// TIA Portal project "Sistema_de_silos" (V16) (continued)
REGION Network 7: Acionamento do Damper / Logica de segurança
   // O ideal é ter o feedback do motor (transportador)
   RUNG wire#powerrail
      Contact( #iCmdAbasteceSilo )
      I_Contact( #iSensorMaximo )
      wire#w1
      Contact( #iSensorDamper01 )
      Contact( #iSensorDamper02 )
      wire#w2
      I_Contact( #Falha_SensoresNivel )
      I_Contact( #Falha_TimeOut_Desabastecimento )
      I_Contact( #iEmg )
      I_Contact( #iCodinicial )
      Coil( #oLigarDumper )
   END_RUNG
   RUNG wire#w1
      Contact( #oLigarDumper )
   END_RUNG wire#w2
   RUNG wire#powerrail
      Contact( #iManual )
      Contact( #btnLigaDumper )
      I_Contact( #"Status Silo - Maximo" )
      Contact( #oLigarTransportador )
      I_Contact( #protecao_damper )
   END_RUNG wire#w2
   // the same network as SCL:
   #oLigarDumper := ((#iCmdAbasteceSilo AND NOT #iSensorMaximo AND ((#iSensorDamper01 AND #iSensorDamper02) OR #oLigarDumper)) OR (#iManual AND #btnLigaDumper AND NOT #"Status Silo - Maximo" AND #oLigarTransportador AND NOT #protecao_damper)) AND NOT #Falha_SensoresNivel AND NOT #Falha_TimeOut_Desabastecimento AND NOT #iEmg AND NOT #iCodinicial;
END_REGION

REGION Network 8: Liga Transportador
   RUNG wire#powerrail
      Contact( #status_damper )
      Contact( #iAutomatico )
      wire#w1
      I_Contact( #Falha_SensoresNivel )
      I_Contact( #Falha_TimeOut_Desabastecimento )
      I_Contact( #iEmg )
      Coil( #oLigarTransportador )
   END_RUNG
   RUNG wire#powerrail
      Contact( #iManual )
      Contact( #btnLigaTransportador )
   END_RUNG wire#w1
   // the same network as SCL:
   #oLigarTransportador := ((#status_damper AND #iAutomatico) OR (#iManual AND #btnLigaTransportador)) AND NOT #Falha_SensoresNivel AND NOT #Falha_TimeOut_Desabastecimento AND NOT #iEmg;
END_REGION

REGION Network 9: Silo Principal - Reserva do produto
   RUNG wire#powerrail
      Contact( #iSensorMinimo )
      wire#w1
      I_Contact( #iSensorMaximo )
      Coil( #"Status Silo - Minimo" )
   END_RUNG
   RUNG wire#w1
      Contact( #iSensorMaximo )
      Coil( #"Status Silo - Maximo" )
   END_RUNG
   RUNG wire#powerrail
      I_Contact( #iSensorMinimo )
      I_Contact( #iSensorMaximo )
      Coil( #"Status Silo - Desabastecido" )
   END_RUNG
   // the same network as SCL:
   #"Status Silo - Minimo" := #iSensorMinimo AND NOT #iSensorMaximo;
   #"Status Silo - Maximo" := #iSensorMinimo AND #iSensorMaximo;
   #"Status Silo - Desabastecido" := NOT #iSensorMinimo AND NOT #iSensorMaximo;
END_REGION

REGION Network 10: Falha dos Sensores de Nivel
   RUNG wire#powerrail
      Contact( #iSensorMaximo )
      I_Contact( #iSensorMinimo )
      S_Coil( #Falha_SensoresNivel )
   END_RUNG
   // the same network as SCL:
   IF #iSensorMaximo AND NOT #iSensorMinimo THEN #Falha_SensoresNivel := TRUE; END_IF;
END_REGION

REGION Network 11: Memoria Auxilar de Erro - Falha de desabastecimento
   RUNG wire#powerrail
      Contact( #"Status Silo - Minimo" )
      Contact( #oAbrirValvula )
      I_Contact( #"Status Silo - Maximo" )
      S_Coil( "DB_Geral".Memoria_Auxiliar_Erro_Silo_1 )
   END_RUNG
   RUNG wire#powerrail
      Contact( #"Status Silo - Desabastecido" )
      R_Coil( "DB_Geral".Memoria_Auxiliar_Erro_Silo_1 )
   END_RUNG
   // the same network as SCL:
   IF #"Status Silo - Minimo" AND #oAbrirValvula AND NOT #"Status Silo - Maximo" THEN
       "DB_Geral".Memoria_Auxiliar_Erro_Silo_1 := TRUE;
   END_IF;
   IF #"Status Silo - Desabastecido" THEN "DB_Geral".Memoria_Auxiliar_Erro_Silo_1 := FALSE; END_IF;
END_REGION

REGION Network 12: Falha de Desabastecimento
   "IEC_Timer_0_DB_TON_TempoErro".TON(IN := "DB_Geral".Memoria_Auxiliar_Erro_Silo_1,
                           PT := "DB_Geral".Time_TempoErro_1);
   IF "IEC_Timer_0_DB_TON_TempoErro".Q THEN #Falha_TimeOut_Desabastecimento := TRUE; END_IF;
END_REGION

REGION Network 13: Reset - Falhas
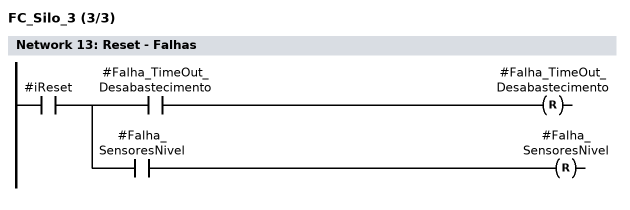
   RUNG wire#powerrail
      Contact( #iReset )
      wire#w1
      Contact( #Falha_TimeOut_Desabastecimento )
      R_Coil( #Falha_TimeOut_Desabastecimento )
   END_RUNG
   RUNG wire#w1
      Contact( #Falha_SensoresNivel )
      R_Coil( #Falha_SensoresNivel )
   END_RUNG
   // the same network as SCL:
   IF #iReset AND #Falha_TimeOut_Desabastecimento THEN #Falha_TimeOut_Desabastecimento := FALSE; END_IF;
   IF #iReset AND #Falha_SensoresNivel THEN #Falha_SensoresNivel := FALSE; END_IF;
END_REGION
END_FUNCTION

FUNCTION "FC_estado_Silos" : Void   // FC8, LAD
{ S7_Optimized_Access := 'TRUE' }
VERSION : 0.1
BEGIN

REGION Network 1
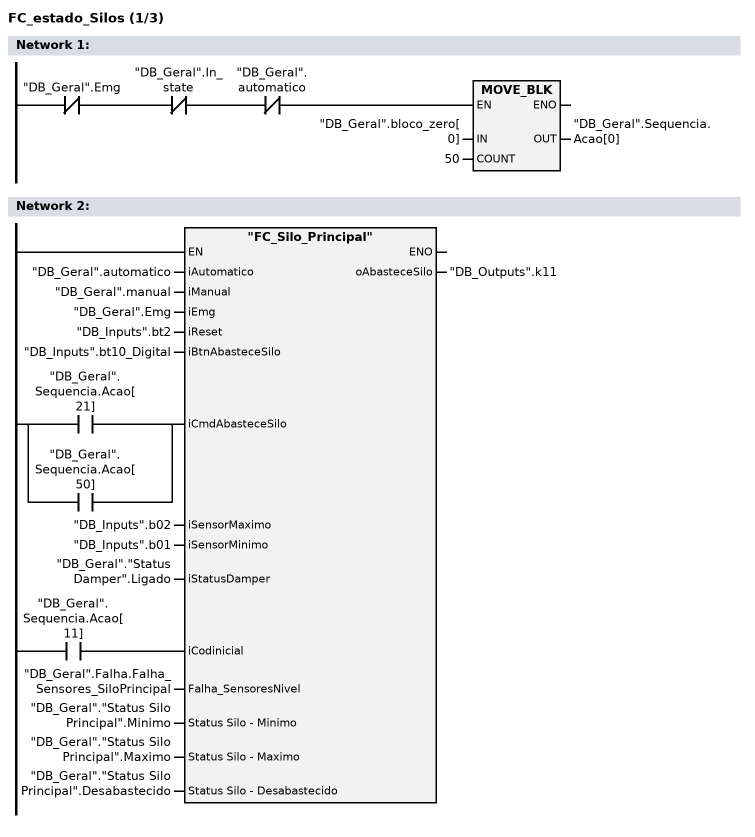
   IF NOT "DB_Geral".Emg AND NOT "DB_Geral".In_state AND NOT "DB_Geral".automatico THEN
       MOVE_BLK(IN := "DB_Geral".bloco_zero[0], COUNT := 50, OUT => "DB_Geral".Sequencia.Acao[0]);
   END_IF;
END_REGION

REGION Network 2
   RUNG wire#powerrail
      "FC_Silo_Principal"(iCmdAbasteceSilo := wire#w1, iCodinicial := wire#w2, iAutomatico := "DB_Geral".automatico, iManual := "DB_Geral".manual, iEmg := "DB_Geral".Emg, iReset := "DB_Inputs".bt2, iBtnAbasteceSilo := "DB_Inputs".bt10_Digital, iSensorMaximo := "DB_Inputs".b02, iSensorMinimo := "DB_Inputs".b01, iStatusDamper := "DB_Geral"."Status Damper".Ligado, Falha_SensoresNivel := "DB_Geral".Falha.Falha_Sensores_SiloPrincipal, "Status Silo - Minimo" := "DB_Geral"."Status Silo Principal".Minimo, "Status Silo - Maximo" := "DB_Geral"."Status Silo Principal".Maximo, "Status Silo - Desabastecido" := "DB_Geral"."Status Silo Principal".Desabastecido, oAbasteceSilo => "DB_Outputs".k11)
   END_RUNG
   RUNG wire#powerrail
      Contact( "DB_Geral".Sequencia.Acao[21] )
   END_RUNG wire#w1
   RUNG wire#powerrail
      Contact( "DB_Geral".Sequencia.Acao[50] )
   END_RUNG wire#w1
   RUNG wire#powerrail
      Contact( "DB_Geral".Sequencia.Acao[11] )
   END_RUNG wire#w2
   // the same network as SCL:
   "FC_Silo_Principal"(iAutomatico := "DB_Geral".automatico,
                       iManual := "DB_Geral".manual,
                       iEmg := "DB_Geral".Emg,
                       iReset := "DB_Inputs".bt2,
                       iBtnAbasteceSilo := "DB_Inputs".bt10_Digital,
                       iCmdAbasteceSilo := "DB_Geral".Sequencia.Acao[21] OR "DB_Geral".Sequencia.Acao[50],
                       iSensorMaximo := "DB_Inputs".b02,
                       iSensorMinimo := "DB_Inputs".b01,
                       iStatusDamper := "DB_Geral"."Status Damper".Ligado,
                       iCodinicial := "DB_Geral".Sequencia.Acao[11],
                       Falha_SensoresNivel := "DB_Geral".Falha.Falha_Sensores_SiloPrincipal,
                       "Status Silo - Minimo" := "DB_Geral"."Status Silo Principal".Minimo,
                       "Status Silo - Maximo" := "DB_Geral"."Status Silo Principal".Maximo,
                       "Status Silo - Desabastecido" := "DB_Geral"."Status Silo Principal".Desabastecido,
                       oAbasteceSilo => "DB_Outputs".k11);
END_REGION

REGION Network 3
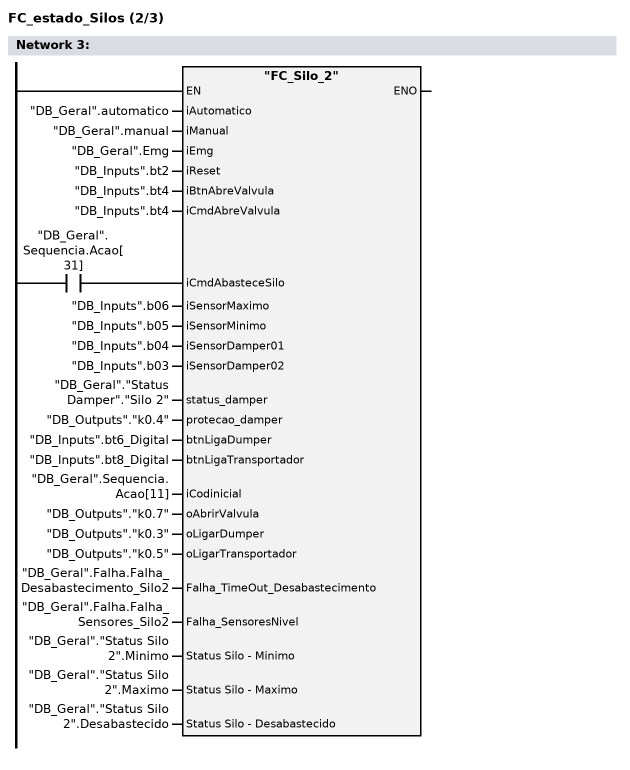
   RUNG wire#powerrail
      "FC_Silo_2"(iCmdAbasteceSilo := wire#w1, iAutomatico := "DB_Geral".automatico, iManual := "DB_Geral".manual, iEmg := "DB_Geral".Emg, iReset := "DB_Inputs".bt2, iBtnAbreValvula := "DB_Inputs".bt4, iCmdAbreValvula := "DB_Inputs".bt4, iSensorMaximo := "DB_Inputs".b06, iSensorMinimo := "DB_Inputs".b05, iSensorDamper01 := "DB_Inputs".b04, iSensorDamper02 := "DB_Inputs".b03, status_damper := "DB_Geral"."Status Damper"."Silo 2", protecao_damper := "DB_Outputs"."k0.4", btnLigaDumper := "DB_Inputs".bt6_Digital, btnLigaTransportador := "DB_Inputs".bt8_Digital, iCodinicial := "DB_Geral".Sequencia.Acao[11], oAbrirValvula := "DB_Outputs"."k0.7", oLigarDumper := "DB_Outputs"."k0.3", oLigarTransportador := "DB_Outputs"."k0.5", Falha_TimeOut_Desabastecimento := "DB_Geral".Falha.Falha_Desabastecimento_Silo2, Falha_SensoresNivel := "DB_Geral".Falha.Falha_Sensores_Silo2, "Status Silo - Minimo" := "DB_Geral"."Status Silo 2".Minimo, "Status Silo - Maximo" := "DB_Geral"."Status Silo 2".Maximo, "Status Silo - Desabastecido" := "DB_Geral"."Status Silo 2".Desabastecido)
   END_RUNG
   RUNG wire#powerrail
      Contact( "DB_Geral".Sequencia.Acao[31] )
   END_RUNG wire#w1
   // the same network as SCL:
   "FC_Silo_2"(iAutomatico := "DB_Geral".automatico,
               iManual := "DB_Geral".manual,
               iEmg := "DB_Geral".Emg,
               iReset := "DB_Inputs".bt2,
               iBtnAbreValvula := "DB_Inputs".bt4,
               iCmdAbreValvula := "DB_Inputs".bt4,
               iCmdAbasteceSilo := "DB_Geral".Sequencia.Acao[31],
               iSensorMaximo := "DB_Inputs".b06,
               iSensorMinimo := "DB_Inputs".b05,
               iSensorDamper01 := "DB_Inputs".b04,
               iSensorDamper02 := "DB_Inputs".b03,
               status_damper := "DB_Geral"."Status Damper"."Silo 2",
               protecao_damper := "DB_Outputs"."k0.4",
               btnLigaDumper := "DB_Inputs".bt6_Digital,
               btnLigaTransportador := "DB_Inputs".bt8_Digital,
               iCodinicial := "DB_Geral".Sequencia.Acao[11],
               oAbrirValvula := "DB_Outputs"."k0.7",
               oLigarDumper := "DB_Outputs"."k0.3",
               oLigarTransportador := "DB_Outputs"."k0.5",
               Falha_TimeOut_Desabastecimento := "DB_Geral".Falha.Falha_Desabastecimento_Silo2,
               Falha_SensoresNivel := "DB_Geral".Falha.Falha_Sensores_Silo2,
               "Status Silo - Minimo" := "DB_Geral"."Status Silo 2".Minimo,
               "Status Silo - Maximo" := "DB_Geral"."Status Silo 2".Maximo,
               "Status Silo - Desabastecido" := "DB_Geral"."Status Silo 2".Desabastecido);
END_REGION

REGION Network 4
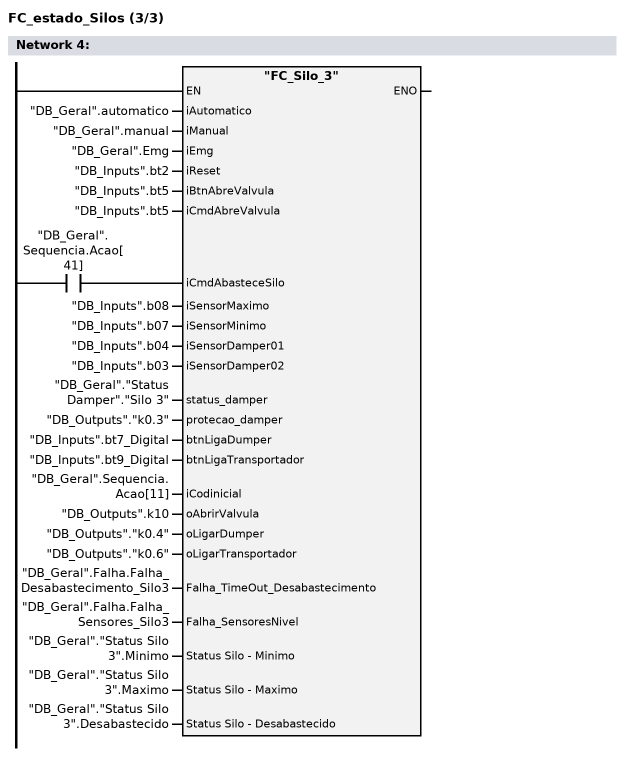
   RUNG wire#powerrail
      "FC_Silo_3"(iCmdAbasteceSilo := wire#w1, iAutomatico := "DB_Geral".automatico, iManual := "DB_Geral".manual, iEmg := "DB_Geral".Emg, iReset := "DB_Inputs".bt2, iBtnAbreValvula := "DB_Inputs".bt5, iCmdAbreValvula := "DB_Inputs".bt5, iSensorMaximo := "DB_Inputs".b08, iSensorMinimo := "DB_Inputs".b07, iSensorDamper01 := "DB_Inputs".b04, iSensorDamper02 := "DB_Inputs".b03, status_damper := "DB_Geral"."Status Damper"."Silo 3", protecao_damper := "DB_Outputs"."k0.3", btnLigaDumper := "DB_Inputs".bt7_Digital, btnLigaTransportador := "DB_Inputs".bt9_Digital, iCodinicial := "DB_Geral".Sequencia.Acao[11], oAbrirValvula := "DB_Outputs".k10, oLigarDumper := "DB_Outputs"."k0.4", oLigarTransportador := "DB_Outputs"."k0.6", Falha_TimeOut_Desabastecimento := "DB_Geral".Falha.Falha_Desabastecimento_Silo3, Falha_SensoresNivel := "DB_Geral".Falha.Falha_Sensores_Silo3, "Status Silo - Minimo" := "DB_Geral"."Status Silo 3".Minimo, "Status Silo - Maximo" := "DB_Geral"."Status Silo 3".Maximo, "Status Silo - Desabastecido" := "DB_Geral"."Status Silo 3".Desabastecido)
   END_RUNG
   RUNG wire#powerrail
      Contact( "DB_Geral".Sequencia.Acao[41] )
   END_RUNG wire#w1
   // the same network as SCL:
   "FC_Silo_3"(iAutomatico := "DB_Geral".automatico,
               iManual := "DB_Geral".manual,
               iEmg := "DB_Geral".Emg,
               iReset := "DB_Inputs".bt2,
               iBtnAbreValvula := "DB_Inputs".bt5,
               iCmdAbreValvula := "DB_Inputs".bt5,
               iCmdAbasteceSilo := "DB_Geral".Sequencia.Acao[41],
               iSensorMaximo := "DB_Inputs".b08,
               iSensorMinimo := "DB_Inputs".b07,
               iSensorDamper01 := "DB_Inputs".b04,
               iSensorDamper02 := "DB_Inputs".b03,
               status_damper := "DB_Geral"."Status Damper"."Silo 3",
               protecao_damper := "DB_Outputs"."k0.3",
               btnLigaDumper := "DB_Inputs".bt7_Digital,
               btnLigaTransportador := "DB_Inputs".bt9_Digital,
               iCodinicial := "DB_Geral".Sequencia.Acao[11],
               oAbrirValvula := "DB_Outputs".k10,
               oLigarDumper := "DB_Outputs"."k0.4",
               oLigarTransportador := "DB_Outputs"."k0.6",
               Falha_TimeOut_Desabastecimento := "DB_Geral".Falha.Falha_Desabastecimento_Silo3,
               Falha_SensoresNivel := "DB_Geral".Falha.Falha_Sensores_Silo3,
               "Status Silo - Minimo" := "DB_Geral"."Status Silo 3".Minimo,
               "Status Silo - Maximo" := "DB_Geral"."Status Silo 3".Maximo,
               "Status Silo - Desabastecido" := "DB_Geral"."Status Silo 3".Desabastecido);
END_REGION
END_FUNCTION

ORGANIZATION_BLOCK "Main"   // OB1, LAD, ProgramCycle
TITLE = "Main Program Sweep (Cycle)"
{ S7_Optimized_Access := 'TRUE' }
VERSION : 0.1
   VAR_INPUT
      Initial_Call : Bool;   // Initial call of this OB
      Remanence : Bool;   // =True, if remanent data are available
   END_VAR
BEGIN

REGION Network 1
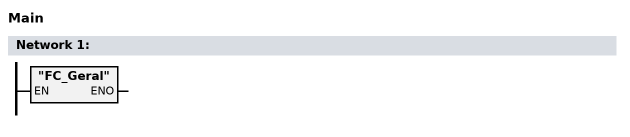
   RUNG wire#powerrail
      "FC_Geral"()
   END_RUNG
   // the same network as SCL:
   "FC_Geral"();
END_REGION
END_ORGANIZATION_BLOCK

(* ===== HMI "HMI_RT_1" =====
system functions are stored by id; their names below are inferred from use
connection "HMI_Connection_2": ETHERNET, S7_1200_OMS

HMI tags "Default tag table"
   "Tag_ScreenNumber" : UInt, internal
   "bt1" : Bool = PLC bt1 AT %I0.1, 1 s
   "bt0" : Bool = PLC bt0 AT %I0.0, 1 s
   "bt3" : Bool = PLC bt3 AT %I0.3, 1 s
   "bt2" : Bool = PLC bt2 AT %I0.2, 1 s
   "DB_Inputs_bt1" : Bool = PLC DB_Inputs.bt1, 1 s
   "DB_Inputs_bt0" : Bool = PLC DB_Inputs.bt0, 1 s
   "DB_Inputs_bt3" : Bool = PLC DB_Inputs.bt3, 1 s
   "DB_Inputs_bt2" : Bool = PLC DB_Inputs.bt2, 1 s
   "DB_Inputs_bt4" : Bool = PLC DB_Inputs.bt4, 1 s
   "DB_Inputs_bt5" : Bool = PLC DB_Inputs.bt5, 1 s
   "DB_Inputs_b04" : Bool = PLC DB_Inputs.b04, 1 s
   "DB_Inputs_b03" : Bool = PLC DB_Inputs.b03, 1 s
   "DB_Outputs_k0.5" : Bool = PLC DB_Outputs."k0.5", 1 s
   "DB_Outputs_k0.6" : Bool = PLC DB_Outputs."k0.6", 1 s
   "DB_Outputs_k0.7" : Bool = PLC DB_Outputs."k0.7", 1 s
   "DB_Geral_Falha_Falha_Desabastecimento_Silo2" : Bool = PLC DB_Geral.Falha.Falha_Desabastecimento_Silo2, 1 s
   "DB_Outputs_k10" : Bool = PLC DB_Outputs.k10, 1 s
   "DB_Geral_Falha_Falha_Desabastecimento_Silo3" : Bool = PLC DB_Geral.Falha.Falha_Desabastecimento_Silo3, 1 s
   "DB_Inputs_b01" : Bool = PLC DB_Inputs.b01, 1 s
   "DB_Geral_Falha_Falha_Sensores_SiloPrincipal" : Bool = PLC DB_Geral.Falha.Falha_Sensores_SiloPrincipal, 1 s
   "DB_Inputs_b02" : Bool = PLC DB_Inputs.b02, 1 s
   "DB_Geral_Falha_Falha_Sensores_Silo2" : Bool = PLC DB_Geral.Falha.Falha_Sensores_Silo2, 1 s
   "DB_Inputs_b05" : Bool = PLC DB_Inputs.b05, 1 s
   "DB_Inputs_b06" : Bool = PLC DB_Inputs.b06, 1 s
   "DB_Geral_Falha_Falha_Sensores_Silo3" : Bool = PLC DB_Geral.Falha.Falha_Sensores_Silo3, 1 s
   "DB_Inputs_b07" : Bool = PLC DB_Inputs.b07, 1 s
   "DB_Inputs_b08" : Bool = PLC DB_Inputs.b08, 1 s
   "DB_Geral_Status Damper_Ligado" : Bool = PLC DB_Geral."Status Damper".Ligado, 1 s
   "DB_Geral_Status Damper_Silo 2" : Bool = PLC DB_Geral."Status Damper"."Silo 2", 1 s
   "DB_Geral_Status Damper_Silo 3" : Bool = PLC DB_Geral."Status Damper"."Silo 3", 1 s
   "DB_Geral_number_status" : Int = PLC DB_Geral.number_status, 1 s
   "DB_Geral_automatico" : Bool = PLC DB_Geral.automatico, 1 s
   "DB_Geral_manual" : Bool = PLC DB_Geral.manual, 1 s
   "DB_Geral_Contador_Abastecimento" : Int = PLC DB_Geral.Contador_Abastecimento, 1 s
   "DB_Outputs_k11" : Bool = PLC DB_Outputs.k11, 1 s
   "DB_Inputs_bt6_Digital" : Bool = PLC DB_Inputs.bt6_Digital, 1 s
   "DB_Inputs_bt7_Digital" : Bool = PLC DB_Inputs.bt7_Digital, 1 s
   "DB_Inputs_bt8_Digital" : Bool = PLC DB_Inputs.bt8_Digital, 1 s
   "DB_Inputs_bt9_Digital" : Bool = PLC DB_Inputs.bt9_Digital, 1 s
   "DB_Inputs_bt10_Digital" : Bool = PLC DB_Inputs.bt10_Digital, 1 s
   "DB_Outputs_x0.0" : Bool = PLC DB_Outputs."x0.0", 1 s
   "DB_Outputs_x0.1" : Bool = PLC DB_Outputs."x0.1", 1 s
   "DB_Outputs_x0.2" : Bool = PLC DB_Outputs."x0.2", 1 s

HMI tags "Animation"
   "Tag_op" : Bool, internal

text list "contador_abastecimento": 0..10000 ''

graphic list "sensor_damper_silo3Aberto": 0 'Group 1000005174'; 1 'sensor_silo3_damper_aberto'

graphic list "sensor_damper_silo2Aberto": 0 'Group 1000005187'; 1 'sensor_silo2_damper_aberto_acionado'

graphic list "transportador": 0 'conveyor'; 1 'transportador_acionado'

graphic list "sensores_nivel": 0 'Sensores_nivel_normal_1'; 1 'sensores_nivel_acionado'

graphic list "valvula2": 0 'valvula2'; 1 'valvula2_acionada'

graphic list "valvula3": 0 'Valvula3'; 1 'Valvula3_acionada'

graphic list "damper": 0 'damper_desligado'

graphic list "damper2": 0 ''; 1 'damper_silo2_acionado'

graphic list "damper3": 0 ''; 1 'damper_silo3_acionado'

graphic list "sensores_nivel_falha": 0 ''; 1 'Sensores_nivel_falha_1'

graphic list "valvula2_Falha": 0 ''; 1 'valvula2_falha'

graphic list "valvula3_falha": 0 ''; 1 'Valvula3_falha'

graphic list "Status": 0 'StatusManual'; 1 'statusAutomatico'; 2 'StatusEmg'; 3 'statusFalha'; 4 'statusSemModo'

graphic list "manual": 0 'StatusManual_off'; 1 'StatusManual'

graphic list "automatico": 0 'statusAutomatico (1)'; 1 'statusAutomatico_1'

graphic list "emergencia": 1 'StatusEmg_off'; 0 'StatusEmg'

graphic list "reset": 0 'statusSemModo_off'; 1 'Reset'

graphic list "btn_valvula2": 0 'Valvula 2 off'; 1 'Valvula 2 ON'

graphic list "btn_valvula3": 0 'Valvula 3 off'; 1 'Valvula 3 ON'

graphic list "AbasteceSiloPrincipal": 0 'Abastece Silo Princiapal_1'; 1 'Abastece Silo Princiapal_on'

graphic list "Btn_damper_s2": 0 'Damper_s2_off'; 1 'Damper_s2ON'

graphic list "Btn_damper_s3": 0 'Damper_s3off'; 1 'Damper_s3ON'

graphic list "btn_transportador1": 0 't1off'; 1 't1ON'

graphic list "btn_transportador2": 0 't2off'; 1 't2ON'

screen "Root screen" 1280x740, template "Template_1"
   on GenerateScreen: SetTag("Tag_ScreenNumber", 1)
   Button "HmiScreenItemData" at 79,35 size 213x73; TextOff 'Teste Screen'; PictureOff "Navigates to Teste Screen for TP1200 Comfort 16.0.0.0"; PictureOn "Navigates to Teste Screen for TP1200 Comfort 16.0.0.0"
      on Release: ActivateScreen("Teste Screen", 0)
   Button "HmiScreenItemData_1" at 1002,36 size 213x73; TextOff 'Operation Screen'; PictureOff "Navigates to Operation Screen for TP1200 Comfort 16.0.0.0"; PictureOn "Navigates to Operation Screen for TP1200 Comfort 16.0.0.0"
      on Release: ActivateScreen("Operation Screen", 0)
   Button "HmiScreenItemData_2" at 692,33 size 213x73; TextOff 'Fail/Emg Screen'; PictureOff "Navigates to Fail/Emg Screen for TP1200 Comfort 16.0.0.0"; PictureOn "Navigates to Fail/Emg Screen for TP1200 Comfort 16.0.0.0"
      on Release: ActivateScreen("Fail/Emg Screen", 0)
   Button "HmiScreenItemData_4" at 377,35 size 213x73; TextOff 'System screens'; PictureOff "Navigates to System screens for TP1200 Comfort 16.0.0.0"; PictureOn "Navigates to System screens for TP1200 Comfort 16.0.0.0"
      on Release: ActivateScreen("System screens", 0)
   GraphicView "Graphic view_3" at 361,257 size 541x174; Picture "Siemens Logo"

Template "Template_1" 1280x740
   Button "Exit" at 1200,679 size 78x59; TextOff 'Exit'; PictureOff "ExitRuntime_TP1200_Comfort_TR"; PictureOn "ExitRuntime_TP1200_Comfort_TR"
      on Release: StopRuntime(0)
   Button "Template_Button" at 1120,679 size 78x59; TextOff 'Text'
   Button "Template_Button_1" at 1040,679 size 78x59; TextOff 'Text'
   Button "Template_Button_2" at 960,679 size 78x59; TextOff 'Text'
   Button "Template_Button_3" at 880,679 size 78x59; TextOff 'Text'
   Button "Template_Button_4" at 800,679 size 78x59; TextOff 'Text'
   Button "Template_Button_5" at 720,679 size 78x59; TextOff 'Text'
   Button "Template_Button_6" at 640,679 size 78x59; TextOff 'Text'
   Button "Template_Button_7" at 561,679 size 78x59; TextOff 'Text'
   Button "Template_Button_8" at 481,679 size 78x59; TextOff 'Text'
   Button "Template_Button_9" at 401,679 size 78x59; TextOff 'Text'
   Button "Template_Button_10" at 321,679 size 78x59; TextOff 'Text'
   Button "Template_Button_11" at 241,679 size 78x59; TextOff 'Text'
   Button "Template_Button_12" at 161,679 size 78x59; TextOff 'Text'
   Button "Alarms" at 81,679 size 78x59; TextOff 'Alarms'; PictureOff "AlarmDisplay_TP1200_Comfort_TR"; PictureOn "AlarmDisplay_TP1200_Comfort_TR"
      on Release: function_ef3f5d25("Alarm window_Unacknowledged", -1)
   Button "Start screen" at 1,679 size 78x59; TextOff 'Start screen'; PictureOff "NavigateHome_TP1200_Comfort_TR"; PictureOn "NavigateHome_TP1200_Comfort_TR"
      on Release: ActivateScreen("Root screen", 0)

screen "Teste Screen" 1280x740, template "Template_1"
   on GenerateScreen: SetTag("Tag_ScreenNumber", 2)
   Rectangle "Rectangle_2" at 211,29 size 201x639
      Visibility <- "Tag_op"
   Rectangle "Rectangle_1" at 0,130 size 201x542
      Visibility <- "Tag_op"
   Button "Back" at 0,0 size 112x36; TextOff 'Back'
      on Release: ActivateScreen("Root screen", 0)
   GraphicView "Graphic view_6" at 768,48 size 165x302; Picture "Clip_path_group_1-removebg-preview"
   Button "Button_5" at 223,153 size 173x77; TextOff 'Text'; PictureOff "btn_val2_1"; PictureList "btn_valvula3"
      Visibility <- "Tag_op"
      on Click: InvertBit("DB_Inputs_bt5")
      ProcessValue <- "DB_Inputs_bt5"
   Button "Button_6" at 224,46 size 173x77; TextOff 'Text'; PictureOff "btn_val3"; PictureList "btn_valvula2"
      Visibility <- "Tag_op"
      on Click: InvertBit("DB_Inputs_bt4")
      ProcessValue <- "DB_Inputs_bt4"
   Button "Button_7" at 0,93 size 199x32; TextOff 'Operação'
      on Click: InvertBit("Tag_op")
   GraphicIOField "Graphic I/O field_1" at 788,246 size 41x16; PictureList "sensor_damper_silo3Aberto"
      ProcessValue <- "DB_Inputs_b04"
   GraphicIOField "Graphic I/O field_2" at 879,245 size 41x16; PictureList "sensor_damper_silo2Aberto"
      ProcessValue <- "DB_Inputs_b03"
   GraphicIOField "Graphic I/O field_3" at 638,372 size 178x32; PictureList "transportador"
      ProcessValue <- "DB_Outputs_k0.5"
   GraphicIOField "Graphic I/O field_4" at 894,371 size 178x32; PictureList "transportador"
      ProcessValue <- "DB_Outputs_k0.6"
   GraphicView "Graphic view_3" at 509,415 size 126x229; Picture "silo2"
   GraphicIOField "Graphic I/O field_5" at 459,623 size 96x20; PictureList "valvula2"
      ProcessValue <- "DB_Outputs_k0.7"
      Visibility <- "DB_Geral_Falha_Falha_Desabastecimento_Silo2"
   GraphicView "Graphic view_5" at 1063,415 size 126x228; Picture "silo2"
   GraphicIOField "Graphic I/O field_6" at 1144,623 size 96x20; PictureList "valvula3"
      ProcessValue <- "DB_Outputs_k10"
      Visibility <- "DB_Geral_Falha_Falha_Desabastecimento_Silo3"
   GraphicIOField "Graphic I/O field_7" at 459,623 size 96x20; PictureList "valvula2_Falha"
      Visibility <- "DB_Geral_Falha_Falha_Desabastecimento_Silo2"
      ProcessValue <- "DB_Geral_Falha_Falha_Desabastecimento_Silo2"
   GraphicIOField "Graphic I/O field_8" at 1144,623 size 96x20; PictureList "valvula3_falha"
      Visibility <- "DB_Geral_Falha_Falha_Desabastecimento_Silo3"
      ProcessValue <- "DB_Geral_Falha_Falha_Desabastecimento_Silo3"
   GraphicIOField "Graphic I/O field_9" at 709,58 size 305x23; PictureList "sensores_nivel"
      Visibility <- "DB_Geral_Falha_Falha_Sensores_SiloPrincipal"
      ProcessValue <- "DB_Inputs_b02"
   GraphicIOField "Graphic I/O field_10" at 712,166 size 305x23; PictureList "sensores_nivel"
      Visibility <- "DB_Geral_Falha_Falha_Sensores_SiloPrincipal"
      ProcessValue <- "DB_Inputs_b01"
   GraphicIOField "Graphic I/O field_13" at 449,519 size 238x23; PictureList "sensores_nivel"
      ProcessValue <- "DB_Inputs_b05"
      Visibility <- "DB_Geral_Falha_Falha_Sensores_Silo2"
   GraphicIOField "Graphic I/O field_14" at 449,519 size 238x23; PictureList "sensores_nivel_falha"
      ProcessValue <- "DB_Geral_Falha_Falha_Sensores_Silo2"
      Visibility <- "DB_Geral_Falha_Falha_Sensores_Silo2"
   GraphicIOField "Graphic I/O field_15" at 449,420 size 238x23; PictureList "sensores_nivel"
      ProcessValue <- "DB_Inputs_b06"
      Visibility <- "DB_Geral_Falha_Falha_Sensores_Silo2"
   GraphicIOField "Graphic I/O field_16" at 449,420 size 238x23; PictureList "sensores_nivel_falha"
      Visibility <- "DB_Geral_Falha_Falha_Sensores_Silo2"
      ProcessValue <- "DB_Geral_Falha_Falha_Sensores_Silo2"
   GraphicIOField "Graphic I/O field_17" at 1008,519 size 238x23; PictureList "sensores_nivel"
      ProcessValue <- "DB_Inputs_b07"
      Visibility <- "DB_Geral_Falha_Falha_Desabastecimento_Silo3"
   GraphicIOField "Graphic I/O field_18" at 1008,519 size 238x23; PictureList "sensores_nivel_falha"
      Visibility <- "DB_Geral_Falha_Falha_Sensores_Silo3"
      ProcessValue <- "DB_Geral_Falha_Falha_Sensores_Silo3"
   GraphicIOField "Graphic I/O field_19" at 1006,420 size 238x23; PictureList "sensores_nivel"
      Visibility <- "DB_Geral_Falha_Falha_Sensores_Silo3"
      ProcessValue <- "DB_Inputs_b08"
   GraphicIOField "Graphic I/O field_20" at 1006,420 size 238x23; PictureList "sensores_nivel_falha"
      ProcessValue <- "DB_Geral_Falha_Falha_Sensores_Silo3"
      Visibility <- "DB_Geral_Falha_Falha_Sensores_Silo3"
   Button "Button_9" at 438,412 size 55x34; TextOff 'Text'
      on Press: InvertBit("DB_Inputs_b06")
   Button "Button_10" at 440,519 size 55x34; TextOff 'Text'
      on Press: InvertBit("DB_Inputs_b05")
   Button "Button_11" at 999,414 size 55x34; TextOff 'Text'
      on Press: InvertBit("DB_Inputs_b08")
   Button "Button_12" at 999,514 size 55x34; TextOff 'Text'
      on Press: InvertBit("DB_Inputs_b07")
   Button "Button_13" at 708,162 size 55x34; TextOff 'Text'
      on Press: InvertBit("DB_Inputs_b01")
   Button "Button_16" at 704,55 size 55x34; TextOff 'Text'
      on Press: InvertBit("DB_Inputs_b02")
   GraphicIOField "Graphic I/O field_21" at 824,247 size 56x54; PictureList "damper3"
      ProcessValue <- "DB_Geral_Status Damper_Silo 3"
      Visibility <- "DB_Geral_Status Damper_Silo 3"
   GraphicIOField "Graphic I/O field_22" at 824,247 size 56x54; PictureList "damper2"
      ProcessValue <- "DB_Geral_Status Damper_Silo 2"
      Visibility <- "DB_Geral_Status Damper_Silo 2"
   GraphicIOField "Graphic I/O field_23" at 824,242 size 60x22; PictureList "damper"
      ProcessValue <- "DB_Geral_Status Damper_Ligado"
      Visibility <- "DB_Geral_Status Damper_Ligado"
   Button "Button_8" at 773,240 size 46x29; TextOff 'Text'
      on Press: InvertBit("DB_Inputs_b04")
   GraphicIOField "Graphic I/O field_12" at 712,166 size 305x23; PictureList "sensores_nivel_falha"
      ProcessValue <- "DB_Geral_Falha_Falha_Sensores_SiloPrincipal"
      Visibility <- "DB_Geral_Falha_Falha_Sensores_SiloPrincipal"
   GraphicIOField "Graphic I/O field_11" at 709,58 size 305x23; PictureList "sensores_nivel_falha"
      Visibility <- "DB_Geral_Falha_Falha_Sensores_SiloPrincipal"
      ProcessValue <- "DB_Geral_Falha_Falha_Sensores_SiloPrincipal"
   Button "Button_1" at 14,145 size 173x77; TextOff 'Text'; PictureOff "StatusManual"; PictureList "manual"
      Visibility <- "Tag_op"
      on Press: InvertBit("DB_Inputs_bt1")
      ProcessValue <- "DB_Inputs_bt1"
   Button "Button_2" at 14,253 size 173x77; TextOff 'Text'; PictureOff "statusAutomatico"; PictureList "automatico"
      Visibility <- "Tag_op"
      on Press: InvertBit("DB_Inputs_bt0")
      ProcessValue <- "DB_Inputs_bt0"
   Button "Button_3" at 14,360 size 173x77; TextOff 'Text'; PictureOff "StatusEmg"; PictureList "emergencia"
      Visibility <- "Tag_op"
      on Press: InvertBit("DB_Inputs_bt3")
      ProcessValue <- "DB_Inputs_bt3"
   Button "Button_4" at 14,468 size 173x77; TextOff 'Text'; PictureOff "Reset"; PictureList "reset"
      Visibility <- "Tag_op"
      on Press: InvertBit("DB_Inputs_bt2")
      ProcessValue <- "DB_Inputs_bt2"
   Button "Button_15" at 223,261 size 173x77; TextOff 'Text'; PictureOff "btn_val2_1"; PictureList "Btn_damper_s2"
      on Click: InvertBit("DB_Inputs_bt6_Digital")
      Visibility <- "Tag_op"
      ProcessValue <- "DB_Inputs_bt6_Digital"
   Button "Button_17" at 223,369 size 173x77; TextOff 'Text'; PictureOff "btn_val2_1"; PictureList "Btn_damper_s3"
      on Click: InvertBit("DB_Inputs_bt7_Digital")
      Visibility <- "Tag_op"
      ProcessValue <- "DB_Inputs_bt7_Digital"
   Button "Button_18" at 223,476 size 173x77; TextOff 'Text'; PictureOff "btn_val2_1"; PictureList "btn_transportador1"
      on Click: InvertBit("DB_Inputs_bt8_Digital")
      Visibility <- "Tag_op"
      ProcessValue <- "DB_Inputs_bt8_Digital"
   Button "Button_19" at 222,577 size 173x77; TextOff 'Text'; PictureOff "btn_val2_1"; PictureList "btn_transportador2"
      on Click: InvertBit("DB_Inputs_bt9_Digital")
      Visibility <- "Tag_op"
      ProcessValue <- "DB_Inputs_bt9_Digital"
   Button "Button_20" at 13,566 size 173x77; TextOff 'Text'; PictureOff "Reset"; PictureList "AbasteceSiloPrincipal"
      on Press: InvertBit("DB_Inputs_bt10_Digital")
      Visibility <- "Tag_op"
      ProcessValue <- "DB_Outputs_k11"
   Button "Button_14" at 879,238 size 46x29; TextOff 'Text'
      on Press: InvertBit("DB_Inputs_b03")

screen "Operation Screen" 1280x740, template "Template_1"
   on GenerateScreen: SetTag("Tag_ScreenNumber", 3)
   TextField "HmiScreenItemData" at 128,324 size 1024x27; Text 'Operation Screen'
   Button "Back" at 1,1 size 159x47; TextOff 'Back'
      on Release: ActivateScreen("Root screen", 0)

screen "Fail/Emg Screen" 1280x740, template "Template_1"
   on GenerateScreen: SetTag("Tag_ScreenNumber", 4)
   TextField "HmiScreenItemData" at 128,324 size 1024x27; Text 'Fail/Emg Screen'
   Button "Back" at 1,1 size 159x47; TextOff 'Back'
      on Release: ActivateScreen("Root screen", 0)

screen "System screens" 1280x740, template "Template_1"
   on GenerateScreen: SetTag("Tag_ScreenNumber", 5)
   Button "Back" at 1,1 size 159x47; TextOff 'Back'
      on Release: ActivateScreen("Root screen", 0)
   Button "HmiScreenItemData" at 36,95 size 159x47; TextOff 'SIMATIC PLC system diagnos...'; PictureOff "Navigates to SIMATIC PLC system diagnostics for TP1200 Comfort 16.0.0.0"; PictureOn "Navigates to SIMATIC PLC system diagnostics for TP1200 Comfort 16.0.0.0"
      on Release: ActivateScreen("SIMATIC PLC system diagnostics", 0)
   Button "HmiScreenItemData_1" at 36,154 size 159x47; TextOff 'System settings'; PictureOff "Navigates to System settings for TP1200 Comfort 16.0.0.0"; PictureOn "Navigates to System settings for TP1200 Comfort 16.0.0.0"
      on Release: ActivateScreen("System settings", 0)
   Button "HmiScreenItemData_2" at 36,213 size 159x47; TextOff 'System information'; PictureOff "Navigates to System information for TP1200 Comfort 16.0.0.0"; PictureOn "Navigates to System information for TP1200 Comfort 16.0.0.0"
      on Release: ActivateScreen("System information", 0)

screen "SIMATIC PLC system diagnostics" 1280x740, template "Template_1"
   on GenerateScreen: SetTag("Tag_ScreenNumber", 6)
   SysDiagControl "HmiScreenItemData" at 1,49 size 1276x623
   Button "Back" at 1,1 size 159x47; TextOff 'Back'
      on Release: ActivateScreen("System screens", 0)

screen "System settings" 1280x740, template "Template_1"
   on GenerateScreen: SetTag("Tag_ScreenNumber", 7)
   Button "Calibrate screen" at 36,95 size 159x47; TextOff 'Calibrate screen'
      on Release: function_bc3e350c()
   Button "Clean screen" at 36,154 size 159x47; TextOff 'Clean screen'
      on Release: function_be740847(30)
   Button "Back" at 1,1 size 159x47; TextOff 'Back'
      on Release: ActivateScreen("System screens", 0)

screen "System information" 1280x740, template "Template_1"
   on GenerateScreen: SetTag("Tag_ScreenNumber", 8)
   TextField "HmiScreenItemData" at 35,51 size 171x28; Text 'HMI device type:'
   TextField "HmiScreenItemData_1" at 241,51 size 1004x28; Text 'TP1200 Comfort 16.0.0.0'
   TextField "HmiScreenItemData_2" at 35,81 size 171x28; Text 'Version:'
   TextField "HmiScreenItemData_3" at 35,111 size 171x28; Text 'Connection:'
   TextField "HmiScreenItemData_4" at 241,111 size 1004x28; Text 'ETHERNET'
   TextField "HmiScreenItemData_5" at 35,141 size 171x28; Text 'PLC:'
   TextField "HmiScreenItemData_6" at 241,141 size 1004x28; Text 'SIMATIC S7 1200'
   Button "Display version" at 241,81 size 1004x28; TextOff 'Display version'
      on Release: function_febcb963(-1)
   Button "Back" at 1,1 size 159x47; TextOff 'Back'
      on Release: ActivateScreen("System screens", 0)
*)